   R509_000_POS : ALIAS FOR R509[0].POS;
   R6 : CONTROL[51];
   R97 : CONTROL[2] := ([0].LEN := 10, [1].LEN := 10);
        [0]   // LEHR SPEED Control word For Lehr Speed averaging Function
        [1]   // LEHR SPEED Control word For lehr Speed standard Deviation
   REL_CRUSH_ALL_OFF : ALIAS FOR I[73].10;
   REL_CRUSH_ALL_ON : ALIAS FOR I[73].11;
   REL_DATARCVD_N : ALIAS FOR O[54].2;
   REL_DATARCVDS : ALIAS FOR O[58].2;
   REL_REJWINLAMPN : ALIAS FOR O[54].3;
   REL_REJWINLAMPS : ALIAS FOR O[58].3;
   Sbr_IN_dCapIndex : DINT; {access Read Only}
   Sbr_IN_dConveyor : DINT; {access Read Only}
   Sbr_IN_dDataLength : DINT; {access Read Only}
   Sbr_IN_DestinationCullet : DINT; {access Read Only}
   Sbr_IN_DestinationID : DINT; {access Read Only}
   Sbr_IN_dIndexHead : DINT; {access Read Only}
   Sbr_IN_dMaskAllowed : DINT; {access Read Only}
   Sbr_IN_Position : DINT; {access Read Only}
   Sbr_IN_PosStart : DINT; {access Read Only}
   Sbr_IN_PosStop : DINT; {access Read Only}
   Sbr_IN_ReasonID : DINT; {access Read Only}
   Sbr_IN_ReentryPosition : DINT; {access Read Only}
   Sbr_IN_ReentryPosition_max : DINT; {access Read Only}
   Sbr_IN_ReentryPosition_min : DINT; {access Read Only}
   Sbr_IN_xHeadPos : BOOL; {access Read Only}
   Sbr_IN_xSendAllCullet : BOOL; {access Read Only}
   Sbr_INO_DestinationLite : DINT; {access Read Only}
   Sbr_INO_tConvoy_SL : UDT_Convoy_SL; {access Read Only}
   Sbr_INO_tConvoyCap_ZC : UDT_ConvoyCap_ZC; {access Read Only}
   Sbr_INO_xALLForDestination : BOOL; {access Read Only}
   Sbr_INO_xAllLiteToCullet : BOOL; {access Read Only}
   Sbr_INO_xAtLeastOneForDestination : BOOL; {access Read Only}
   Sbr_INO_xAtLeastOneToCullet : BOOL; {access Read Only}
   Sbr_OUT_dIndexTail : DINT; {access Read Only}
   Sbr_OUT_dTotalCaps : DINT; {access Read Only}
   Sbr_OUT_ReqRot_CCW : BOOL; {access Read Only}
   Sbr_OUT_ReqRot_CW : BOOL; {access Read Only}
   Sbr_OUT_rgdConvoyGaps : DINT[4]; {access Read Only}
   Sbr_OUT_rgdConvoyLengths : DINT[4]; {access Read Only}
   SLOW_BLINK : ALIAS FOR T4[0];
   Speed_Offset_CM07N : DINT := -20;   // This was added to allow for speed adjustment to CM07N
   Speed_Offset_Result_CM07N : DINT := 237;
   T103 : TIMER[1];
   T108 : TIMER[1];
   T113 : TIMER[1];
   T118 : TIMER[1];
   T123 : TIMER[1];
   T128 : TIMER[1];
   T133 : TIMER[1];
   T182 : TIMER[11] := ([0].PRE := 5, [0].ACC := 5, [0].EN := 1, [0].DN := 1, [1].PRE := 50, [2].PRE := 1, [2].ACC := 3, [2].EN := 1, [2].DN := 1, [3].PRE := 30, [4].PRE := 10, [5].PRE := 20000, [5].ACC := 25, [5].EN := 1, [5].TT := 1, [6].PRE := 100, [7].PRE := 500, [8].PRE := 500, [8].ACC := 201, [8].EN := 1, [8].TT := 1, [9].PRE := 10, [10].PRE := 100);
        [7]   // VMCC M2 Speed zone 2 Start Test Timer * M2CM2
        [8]   // VMCC M2 Speed zone 2 Stop Test Timer * M2CM2
   T4 : TIMER[51] := ([0].PRE := 1000, [0].ACC := 220, [0].EN := 1, [0].TT := 1, [1].PRE := 1000, [2].PRE := 500, [3].PRE := 500, [4].PRE := 10000, [8].PRE := 200, [9].PRE := 500, [10].PRE := 500, [11].PRE := 60, [13].PRE := 60000, [13].ACC := 60002, [13].EN := 1, [13].DN := 1, [26].PRE := 2500, [27].PRE := 2500, [28].PRE := 2500, [29].PRE := 2500, [30].PRE := 12000, [30].ACC := 12001, [30].EN := 1, [30].DN := 1, [31].PRE := 100, [31].ACC := 101, [31].EN := 1, [31].DN := 1, [33].PRE := 2500, [34].PRE := 2500, [35].PRE := 2500, [36].PRE := 2500, [37].PRE := 2500, [38].PRE := 2500, [39].PRE := 2500, [40].PRE := 2500, [41].PRE := 2500, [42].PRE := 2500, [43].PRE := 2500, [44].PRE := 2500, [45].PRE := 2500, [46].PRE := 2500, [47].PRE := 2500, [48].PRE := 2500, [49].PRE := 2500, [50].PRE := 2500);
        [0]   // Slow blink On time Timer
        [44]   // M2CM09N Running Delay Timer
        [31]   // M2CMO2 Stopped Failure Detect Debounce timer
        [43]   // M2CM09S Running Delay Timer
        [42]   // M2CM08N Running Delay Timer
        [1]   // Slow blink off time timer
        [26]   // M2CM01 Running Delay Timer
        [29]   // M2CM04S Running Delay Timer
        [2]   // Fast blink On time timer
        [28]   // M2CM03 Running Delay Timer
        [3]   // Fast Blink off time timer
        [39]   // M2CM07S Running Delay Timer
        [8]   // Conv 12 drive enable timer
        [27]   // M2CM02 Running Delay Timer
        [34]   // M2CM04N Running Delay Timer
        [35]   // M2CM05S Running Delay Timer
        [38]   // M2CM06N Running Delay Timer
        [33]   // VMCC M2 Drive Fault timer hold to see if fault will clear
        [37]   // M2CM06S Running Delay Timer
        [36]   // M2CM05N Running Delay Timer
        [40]   // M2CM07N Running Delay Timer
        [41]   // M2CM08S Running Delay Timer
        [46]   // M2CM10N Running Delay Timer
        [47]   // M2CM11S Running Delay Timer
        [48]   // M2CM011N Running Delay Timer
        [49]   // M2CM012S Running Delay Timer
        [30]   // Drive Stopped Failure Detect Debounce timer (All drives were running prev)
        [13]   // BENCHBOARD Timer for CROSSBREAK ON duration (60 sec.)
        [11]   // Test Timer
        [4]   // M4-->>M2 Mainline Sec. Trans. Backup delay timer
        [50]   // M2CM012N Running Delay Timer
        [45]   // M2CM10S Running Delay Timer
   T47 : TIMER[32];
        [10]   // Conveyor 10 Resync Input Debounce Timer
        [11]   // Conveyor 11 Resync Input Debounce Timer
        [12]   // Conveyor 12 Resync Input Debounce Timer
        [19]   // Conveyor 19 Resync Input Debounce Timer
        [1]   // Conveyor 1 Resync Input Debounce Timer
        [20]   // Conveyor 20 Resync Input Debounce Timer
        [21]   // Conveyor 21 Resync Input Debounce Timer
        [22]   // Conveyor 22 Resync Input Debounce Timer
        [23]   // Conveyor 23 Resync Input Debounce Timer
        [24]   // Conveyor 24 Resync Input Debounce Timer
        [25]   // Conveyor 25 Resync Input Debounce Timer
        [26]   // Conveyor 26 Resync Input Debounce Timer
        [27]   // Conveyor 27 Resync Input Debounce Timer
        [28]   // Conveyor 28 Resync Input Debounce Timer
        [29]   // Conveyor 29 Resync Input Debounce Timer
        [2]   // Conveyor 2 Resync Input Debounce Timer
        [30]   // Conveyor 30 Resync Input Debounce Timer
        [31]   // Conveyor 31 Resync Input Debounce Timer
        [13]   // Conveyor 13 Resync Input Debounce Timer
        [3]   // Conveyor 3 Resync Input Debounce Timer
        [4]   // Conveyor 4 Resync Input Debounce Timer
        [5]   // Conveyor 5 Resync Input Debounce Timer
        [6]   // Conveyor 6 Resync Input Debounce Timer
        [7]   // Conveyor 7 Resync Input Debounce Timer
        [8]   // Conveyor 8 Resync Input Debounce Timer
        [9]   // Conveyor 9 Resync Input Debounce Timer
        [14]   // Conveyor 14 Resync Input Debounce Timer
        [15]   // Conveyor 15 Resync Input Debounce Timer
        [16]   // Conveyor 16 Resync Input Debounce Timer
        [17]   // Conveyor 17 Resync Input Debounce Timer
        [18]   // Conveyor 18 Resync Input Debounce Timer
   T9 : TIMER[22] := ([10].PRE := 8000, [10].ACC := 8002, [10].EN := 1, [10].DN := 1, [11].PRE := 8000, [11].ACC := 8001, [11].EN := 1, [11].DN := 1, [12].PRE := 8000, [12].ACC := 8001, [12].EN := 1, [12].DN := 1, [13].PRE := 8000, [13].ACC := 8002, [13].EN := 1, [13].DN := 1, [14].PRE := 8000, [14].ACC := 8001, [14].EN := 1, [14].DN := 1, [15].PRE := 8000, [15].ACC := 8000, [15].EN := 1, [15].DN := 1, [16].PRE := 8000, [16].ACC := 8002, [16].EN := 1, [16].DN := 1, [17].PRE := 8000, [17].ACC := 8002, [17].EN := 1, [17].DN := 1, [18].PRE := 8000, [18].ACC := 8001, [18].EN := 1, [18].DN := 1, [19].PRE := 8000, [19].ACC := 8000, [19].EN := 1, [19].DN := 1, [20].PRE := 8000, [20].ACC := 8001, [20].EN := 1, [20].DN := 1, [21].PRE := 8000, [21].ACC := 8001, [21].EN := 1, [21].DN := 1);
        [10]   // Conv 1 drive enable timer
        [11]   // Conv 2 drive enable timer
        [12]   // Conv 3 drive enable timer
        [13]   // Conv 4 drive enable timer
        [14]   // Conv 5 drive enable timer
        [15]   // Conv 6 drive enable timer
        [16]   // Conv 7 drive enable timer
        [17]   // Conv 8 drive enable timer
        [18]   // Conv 9 drive enable timer
        [19]   // Conv 10 drive enable timer
        [20]   // Conv 11 drive enable timer
        [21]   // Conv 12 drive enable timer
   T95 : TIMER[10] := ([0].PRE := 1000);
        [0].DN   // LEHR SPEED Sample Period timer Elapsed
        [0]   // LEHR SPEED Sample period Timer
   TD1_N_MOVIN : ALIAS FOR N14[256].2;
   TD1_N_MOVOUT : ALIAS FOR N14[257].2;
   TD1_S_MOVIN : ALIAS FOR N14[256].3;
   TD1_S_MOVOUT : ALIAS FOR N14[257].3;
   TD2_N_MOVIN : ALIAS FOR N14[256].4;
   TD2_N_MOVOUT : ALIAS FOR N14[257].4;
   TD2_S_MOVIN : ALIAS FOR N14[256].5;
   TD2_S_MOVOUT : ALIAS FOR N14[257].5;
   TD3_N_MOVIN : ALIAS FOR N14[256].6;
   TD3_N_MOVOUT : ALIAS FOR N14[257].6;
   TD3_S_MOVIN : ALIAS FOR N14[256].7;
   TD3_S_MOVOUT : ALIAS FOR N14[257].7;
   TD4_N_MOVIN : ALIAS FOR N14[256].8;
   TD4_N_MOVOUT : ALIAS FOR N14[257].8;
   TD4_S_MOVIN : ALIAS FOR N14[256].9;
   TD4_S_MOVOUT : ALIAS FOR N14[257].9;
   TD5_N_MOVIN : ALIAS FOR N14[256].10;
   TD5_N_MOVOUT : ALIAS FOR N14[257].10;
   TD5_S_MOVIN : ALIAS FOR N14[256].11;
   TD5_S_MOVOUT : ALIAS FOR N14[257].11;
   TD_ALM_HORN_RLY : ALIAS FOR O[21].3;
   TD_ALM_LAMP : ALIAS FOR I[18].4;
   TD_ALM_RESET : ALIAS FOR I[17].9;
   TD_ALM_SILENCE : ALIAS FOR I[17].8;
   TD_AMBER_STKLTE : ALIAS FOR O[21].6;
   TD_BLUE_STKLTE : ALIAS FOR O[21].5;
   TD_CS2S_Crush_All_Stacklight : ALIAS FOR O[70].15;   // Red Light mounted on the top of panel
   TD_DC_INPWR : ALIAS FOR I[17].2;
   TD_DC_OUTPWR : ALIAS FOR I[17].3;
   TD_DC_PS1 : ALIAS FOR I[17].4;
   TD_DC_PS2 : ALIAS FOR I[17].6;
   TD_DC_PS3 : ALIAS FOR I[17].7;
   TD_DRV_CONT_ON : ALIAS FOR I[17].1;
   TD_DRV_FLT_LMP : ALIAS FOR O[21].0;
   TD_ESTOP : ALIAS FOR I[17].10;
   TD_ESTOPPWR : ALIAS FOR I[17].5;
   TD_FLT_RES_RLY : ALIAS FOR O[21].1;
   TD_RED_STKLTE : ALIAS FOR O[21].4;
   TDN_CRUSH_ALL_OFF : ALIAS FOR I[44].12;
   TDN_CRUSH_ALL_ON : ALIAS FOR I[44].13;
   TDN_FLT : ALIAS FOR I[18].1;
   TDN_FWD : ALIAS FOR O[20].1;
   TDN_REV : ALIAS FOR O[20].5;
   TDN_SS1 : ALIAS FOR O[20].13;
   TDN_SS2 : ALIAS FOR O[20].9;
   TDS_CRUSH_ALL_OFF : ALIAS FOR I[64].12;
   TDS_CRUSH_ALL_ON : ALIAS FOR I[64].13;
   TDS_FLT : ALIAS FOR I[18].2;
   TDS_FWD : ALIAS FOR O[20].2;
   TDS_REV : ALIAS FOR O[20].6;
   TDS_SS1 : ALIAS FOR O[20].14;
   TDS_SS2 : ALIAS FOR O[20].10;
   TEST_OPERAND : ALIAS FOR N7[11];
   TEST_TIMER : ALIAS FOR T4[11];
   TK1_N_MOVDN : ALIAS FOR N14[253].2;
   TK1_N_MOVIN : ALIAS FOR N14[254].2;
   TK1_N_MOVOUT : ALIAS FOR N14[255].2;
   TK1_N_MOVUP : ALIAS FOR N14[252].2;
   TK1_S_MOVDN : ALIAS FOR N14[253].3;
   TK1_S_MOVIN : ALIAS FOR N14[254].3;
   TK1_S_MOVOUT : ALIAS FOR N14[255].3;
   TK1_S_MOVUP : ALIAS FOR N14[252].3;
   TK2_N_MOVDN : ALIAS FOR N14[253].4;
   TK2_N_MOVIN : ALIAS FOR N14[254].4;
   TK2_N_MOVOUT : ALIAS FOR N14[255].4;
   TK2_N_MOVUP : ALIAS FOR N14[252].4;
   TK2_S_MOVDN : ALIAS FOR N14[253].5;
   TK2_S_MOVIN : ALIAS FOR N14[254].5;
   TK2_S_MOVOUT : ALIAS FOR N14[255].5;
   TK2_S_MOVUP : ALIAS FOR N14[252].5;
   TK3_N_MOVDN : ALIAS FOR N14[253].6;
   TK3_N_MOVIN : ALIAS FOR N14[254].6;
   TK3_N_MOVOUT : ALIAS FOR N14[255].6;
   TK3_N_MOVUP : ALIAS FOR N14[252].6;
   TK3_S_MOVDN : ALIAS FOR N14[253].7;
   TK3_S_MOVIN : ALIAS FOR N14[254].7;
   TK3_S_MOVOUT : ALIAS FOR N14[255].7;
   TK3_S_MOVUP : ALIAS FOR N14[252].7;
   TK4_N_MOVDN : ALIAS FOR N14[253].8;
   TK4_N_MOVIN : ALIAS FOR N14[254].8;
   TK4_N_MOVOUT : ALIAS FOR N14[255].8;
   TK4_N_MOVUP : ALIAS FOR N14[252].8;
   TK4_S_MOVDN : ALIAS FOR N14[253].9;
   TK4_S_MOVIN : ALIAS FOR N14[254].9;
   TK4_S_MOVOUT : ALIAS FOR N14[255].9;
   TK4_S_MOVUP : ALIAS FOR N14[252].9;
   TK5_N_MOVDN : ALIAS FOR N14[253].10;
   TK5_N_MOVIN : ALIAS FOR N14[254].10;
   TK5_N_MOVOUT : ALIAS FOR N14[255].10;
   TK5_N_MOVUP : ALIAS FOR N14[252].10;
   TK5_S_MOVDN : ALIAS FOR N14[253].11;
   TK5_S_MOVIN : ALIAS FOR N14[254].11;
   TK5_S_MOVOUT : ALIAS FOR N14[255].11;
   TK5_S_MOVUP : ALIAS FOR N14[252].11;
   TK_FLT : ALIAS FOR I[18].0;
   TK_FWD : ALIAS FOR O[20].0;
   TK_REV : ALIAS FOR O[20].4;
   TK_SS1 : ALIAS FOR O[20].12;
   TK_SS2 : ALIAS FOR O[20].8;
   TMP_CenterLites : BOOL; {access Read Only}
   TMP_d : DINT; {access Read Only}
   TMP_d2 : DINT; {access Read Only}
   TMP_dAccSpace : DINT; {access Read Only}
   TMP_dActualOnLHS : DINT; {access Read Only}
   TMP_dActualSpeed : DINT; {access Read Only}
   TMP_dALARM_RT999 : DINT := 9999; {access None}
   TMP_dBaryc_ins_max : DINT; {access Read Only}
   TMP_dBaryc_ins_min : DINT; {access Read Only}
   TMP_dBufferIndex : DINT; {access Read Only}
   TMP_dBufferSize : DINT; {access Read Only}
   TMP_dCap : DINT; {access Read Only}
   TMP_dCapNextConvoy : DINT; {access Read Only}
   TMP_dConv : DINT; {access Read Only}
   TMP_dConvDebug : DINT; {access Read Only}
   TMP_dConveyorLength : DINT; {access Read Only}
   TMP_dConveyorNumberForZoneCleaning : DINT; {access Read Only}
   TMP_dConvoySearchMax : DINT; {access Read Only}
   TMP_dCountDest : DINT; {access Read Only}
   TMP_dCulletMask : DINT; {access Read Only}
   TMP_dDebug : DINT; {access Read Only}
   TMP_dDecelerationPositionEndConveyor : DINT; {access Read Only}
   TMP_dDecSpace : DINT; {access Read Only}
   TMP_dDestFile : DINT := 205; {access None}
   TMP_dDestOffset : DINT := 1; {access None}
   TMP_dDiffPhotocellStartConv0 : DINT; {access Read Only}
   TMP_dDirection : DINT; {access None}
   TMP_dEndConveyorPos : DINT; {access Read Only}
   TMP_dEndSearch0 : DINT; {access Read Only}
   TMP_dEndSearch1 : DINT; {access Read Only}
   TMP_dErrDestFile : DINT; {access None}
   TMP_dErrSourceFile : DINT; {access None}
   TMP_dFixedSideOffset : DINT; {access Read Only}
   TMP_dFixedSideOffsetBoth : DINT; {access Read Only}
   TMP_dFixedSideOffsetConvoy : DINT; {access Read Only}
   TMP_dFixedSideOffsetDW : DINT; {access Read Only}
   TMP_dFixedSideOffsetUP : DINT; {access Read Only}
   TMP_dHalfConveyorLength : DINT; {access Read Only}
   TMP_dHalfPlateLength : DINT; {access Read Only}
   TMP_dHalfWidthDifference : DINT; {access Read Only}
   TMP_dHeadMax : DINT; {access Read Only}
   TMP_dHeadPosition : DINT; {access Read Only}
   TMP_dHeadPosition_mm : DINT; {access Read Only}
   TMP_dIndC : DINT; {access Read Only}
   TMP_dIndex : DINT := 200;
   TMP_dIndex2 : DINT; {access Read Only}
   TMP_dIndex3 : DINT; {access Read Only}
   TMP_dIndex4 : DINT; {access Read Only}
   TMP_dIndexCap : DINT; {access Read Only}
   TMP_dIndexCapConv : DINT; {access Read Only}
   TMP_dIndexConv : DINT; {access Read Only}
   TMP_dIndexMotor : DINT; {access Read Only}
   TMP_dIndexNext : DINT; {access Read Only}
   TMP_dIndexNextDebug : DINT; {access Read Only}
   TMP_dIndexPlate : DINT; {access Read Only}
   TMP_dIndexPrevious : DINT; {access Read Only}
   TMP_dIndexPreviousDebug : DINT; {access Read Only}
   TMP_DistanceLateralSquaringToCenter : DINT; {access Read Only}
   TMP_dLastConv : DINT; {access Read Only}
   TMP_dLastConvTail : DINT; {access Read Only}
   TMP_dLehrSpeed : DINT; {access Read Only}
   TMP_dLineSize : DINT; {access Read Only}
   TMP_dLineSpeed : DINT; {access Read Only}
   TMP_dLite : DINT; {access Read Only}
   TMP_dLiteInv : DINT; {access Read Only}
   TMP_dManualTargetPos : DINT; {access Read Only}
   TMP_dMask : DINT; {access Read Only}
   TMP_dMaskAllowed : DINT; {access Read Only}
   TMP_dMaxCap : DINT; {access Read Only}
   TMP_dMaxLite : DINT; {access Read Only}
   TMP_dMinTail : DINT; {access Read Only}
   TMP_dMissingOnLHS : DINT; {access Read Only}
   TMP_dNextCap : DINT; {access Read Only}
   TMP_dNumFile : DINT := 648; {access None}
   TMP_dNumValues : DINT := 99; {access None}
   TMP_dOffset : DINT := 32; {access None}
   TMP_dOffsetLoadUnload_cmm : DINT; {access Read Only}
   TMP_dPhEndPosition_cmm : DINT; {access Read Only}
   TMP_dPointer : DINT; {access Read Only}
   TMP_dPointerCap : DINT; {access Read Only}
   TMP_dPos_cmm : DINT; {access Read Only}
   TMP_dPosHead_cmm : DINT; {access Read Only}
   TMP_dPosTail_cmm : DINT; {access Read Only}
   TMP_dRampMotor : DINT; {access Read Only}
   TMP_dSourceFile : DINT := 200; {access None}
   TMP_dSourceOffset : DINT; {access None}
   TMP_dStart0 : DINT; {access Read Only}
   TMP_dStart1 : DINT; {access Read Only}
   TMP_dStartSearch : DINT; {access Read Only}
   TMP_dStartSearch0 : DINT; {access Read Only}
   TMP_dStartSearch1 : DINT; {access Read Only}
   TMP_dStartSearchStop : DINT; {access Read Only}
   TMP_dStepAdvMotor : DINT; {access Read Only}
   TMP_dStop0 : DINT; {access Read Only}
   TMP_dStop1 : DINT; {access Read Only}
   TMP_dStopSearch : DINT; {access Read Only}
   TMP_dStopSearchStop : DINT; {access Read Only}
   TMP_dTailOnNextConveyor_cmm : DINT; {access Read Only}
   TMP_dTailPosition : DINT; {access Read Only}
   TMP_dTarget : DINT := 1815; {access None}
   TMP_dTotalLength : DINT; {access Read Only}
   TMP_dWander : DINT; {access Read Only}
   TMP_dWidth_mm : DINT; {access Read Only}
   TMP_HeadPos : DINT; {access Read Only}
   TMP_IdxLite : DINT; {access Read Only}
   TMP_LiteAHeadY : DINT; {access Read Only}
   TMP_LiteATailY : DINT; {access Read Only}
   TMP_LiteBHeadY : DINT; {access Read Only}
   TMP_LiteBTailY : DINT; {access Read Only}
   TMP_MOV_dDestinationVar_1 : DINT := 205; {access None}
   TMP_MOV_dDestinationVar_2 : DINT; {access None}
   TMP_MOV_dSource : DINT; {access None}
   TMP_OUT_xPlateEndTracking : BOOL; {access Read Only}
   TMP_Portrait : BOOL; {access Read Only}
   TMP_r : REAL; {access Read Only}
   TMP_r1 : REAL := 1900.0; {access None}
   TMP_rAcc : REAL := 1200.0; {access None}
   TMP_rActualValue_cmm : REAL; {access Read Only}
   TMP_rDec : REAL := 1200.0; {access None}
   TMP_rgdIndexC : DINT[4] := ([0] := 2); {access None}
   TMP_rgdPnt : DINT[5]; {access Read Only}
   TMP_rgxId : DINT[10]; {access Read Only}
   TMP_rSpeed : REAL := 1500.0; {access None}
   TMP_rTarget : REAL; {access Read Only}
   TMP_rTarget_M1 : REAL; {access Read Only}
   TMP_rTarget_M2 : REAL; {access Read Only}
   TMP_rTarget_M3 : REAL; {access Read Only}
   TMP_SendToCullet : BOOL; {access Read Only}
   TMP_SquaringPosition : DINT; {access Read Only}
   TMP_StartPlusLength : DINT; {access Read Only}
   TMP_string : STRING; {access Read Only}
   TMP_x : BOOL; {access Read Only}
   TMP_xAllCullet : BOOL; {access Read Only}
   TMP_xALLForSideLeg : BOOL; {access Read Only}
   TMP_xAllLiteToCullet : BOOL; {access Read Only}
   TMP_xAlwaysOFF : BOOL; {access Read Only}
   TMP_xAtLeastOneForQuality : BOOL; {access Read Only}
   TMP_xAtLeastOneForSideLeg : BOOL; {access Read Only}
   TMP_xAtLeastOneOK : BOOL; {access Read Only}
   TMP_xAtLeastOneToCullet : BOOL; {access Read Only}
   TMP_xCenterFound : BOOL; {access Read Only}
   TMP_xConveyorInvolvedInCleaning : BOOL; {access Read Only}
   TMP_xConveyorOfStartCleaning : BOOL; {access Read Only}
   TMP_xCulletPresent : BOOL; {access Read Only}
   TMP_xDebugOFF : BOOL; {access Read Only}
   TMP_xDebugON : BOOL := 1; {access Read Only}
   TMP_xDummy : BOOL; {access Read Only}
   TMP_xEnableLoadUnload : BOOL; {access Read Only}
   TMP_xEnableZoneCleaning : BOOL; {access Read Only}
   TMP_xFirstConv : BOOL; {access Read Only}
   TMP_xForwardCommadnForCleaningZone : BOOL; {access Read Only}
   TMP_xInitialize : BOOL; {access None}
   TMP_xJustOnePlateMissing : BOOL; {access Read Only}
   TMP_xLastConv : BOOL; {access Read Only}
   TMP_xLastConvDebug : BOOL; {access Read Only}
   TMP_xLastModalityLoadBwd : BOOL; {access Read Only}
   TMP_xLastModalityUnloadBwd : BOOL; {access Read Only}
   TMP_xLiteThisDestPresent : BOOL; {access Read Only}
   TMP_xMinTailFound : BOOL; {access Read Only}
   TMP_xOSN : DINT; {access None}
   TMP_xOSN_B : DINT; {access Read Only}
   TMP_xOSR : DINT; {access None}
   TMP_xOSR_B : DINT; {access Read Only}
   TMP_xOSRDebug : BOOL := 1; {access Read Only}
   TMP_xPlateFound : BOOL; {access Read Only}
   TMP_xPlateOnConvoyOnNextConveyor : BOOL; {access Read Only}
   TMP_xPosHead : BOOL; {access Read Only}
   TMP_xPositioning : BOOL; {access Read Only}
   TMP_xPositioning_M1 : BOOL; {access Read Only}
   TMP_xPositioning_M2 : BOOL; {access Read Only}
   TMP_xPositioning_M3 : BOOL; {access Read Only}
   TMP_xPowerSaving : BOOL; {access Read Only}
   TMP_xPresenceAlternative : BOOL; {access Read Only}
   TMP_xPresenceDestination : BOOL; {access Read Only}
   TMP_xPresenceSecondDestination : BOOL; {access Read Only}
   TMP_xReqStopM310M1 : BOOL; {access Read Only}
   TMP_xReqStopM310M2 : BOOL; {access Read Only}
   TMP_xReqStopM310M3 : BOOL; {access Read Only}
   TMP_xReqStopM315M1 : BOOL; {access Read Only}
   TMP_xReqStopM315M2 : BOOL; {access Read Only}
   TMP_xReqStopM315M3 : BOOL; {access Read Only}
   TMP_xReqUnpack : BOOL; {access Read Only}
   TMP_xReverse : BOOL; {access Read Only}
   TMP_xReverse_M1 : BOOL; {access Read Only}
   TMP_xReverse_M2 : BOOL; {access Read Only}
   TMP_xReverse_M3 : BOOL; {access Read Only}
   TMP_xRun : BOOL; {access Read Only}
   TMP_xRun_M1 : BOOL; {access Read Only}
   TMP_xRun_M2 : BOOL; {access Read Only}
   TMP_xRun_M3 : BOOL; {access Read Only}
   TMP_xSimulationActive : BOOL; {access Read Only}
   TMP_xTailFound : BOOL; {access Read Only}
   TMP_xYInversionLite : BOOL; {access Read Only}
   TMP_xYWithBarycenter : BOOL; {access Read Only}
   TMR_Power_Cycle : TIMER := (PRE := 1000, ACC := 1001, EN := 1, DN := 1);
   tony_always_false : BOOL; {access Read Only}
   TRIM_SPEED : ALIAS FOR N20[2];
   TZ1_K_NTH_ADJ : ALIAS FOR O[19].2;
   TZ1_K_STH_ADJ : ALIAS FOR O[19].3;
   TZ1_N_AUTO : ALIAS FOR N14[250].2;
   TZ1_N_MANL : ALIAS FOR N14[251].2;
   TZ1_S_AUTO : ALIAS FOR N14[250].3;
   TZ1_S_MANL : ALIAS FOR N14[251].3;
   TZ1_T_NTH_ADJ : ALIAS FOR O[22].2;
   TZ1_T_STH_ADJ : ALIAS FOR O[22].3;
   TZ2_K_NTH_ADJ : ALIAS FOR O[19].4;
   TZ2_K_STH_ADJ : ALIAS FOR O[19].5;
   TZ2_N_AUTO : ALIAS FOR N14[250].4;
   TZ2_N_MANL : ALIAS FOR N14[251].4;
   TZ2_S_AUTO : ALIAS FOR N14[250].5;
   TZ2_S_MANL : ALIAS FOR N14[251].5;
   TZ2_T_NTH_ADJ : ALIAS FOR O[22].4;
   TZ2_T_STH_ADJ : ALIAS FOR O[22].5;
   TZ3_K_NTH_ADJ : ALIAS FOR O[19].6;
   TZ3_K_STH_ADJ : ALIAS FOR O[19].7;
   TZ3_N_AUTO : ALIAS FOR N14[250].6;
   TZ3_N_MANL : ALIAS FOR N14[251].6;
   TZ3_S_AUTO : ALIAS FOR N14[250].7;
   TZ3_S_MANL : ALIAS FOR N14[251].7;
   TZ3_T_NTH_ADJ : ALIAS FOR O[22].6;
   TZ3_T_STH_ADJ : ALIAS FOR O[22].7;
   TZ4_K_NTH_ADJ : ALIAS FOR O[19].8;
   TZ4_K_STH_ADJ : ALIAS FOR O[19].9;
   TZ4_N_AUTO : ALIAS FOR N14[250].8;
   TZ4_N_MANL : ALIAS FOR N14[251].8;
   TZ4_S_AUTO : ALIAS FOR N14[250].9;
   TZ4_S_MANL : ALIAS FOR N14[251].9;
   TZ4_T_NTH_ADJ : ALIAS FOR O[22].8;
   TZ4_T_STH_ADJ : ALIAS FOR O[22].9;
   TZ5_K_NTH_ADJ : ALIAS FOR O[19].10;
   TZ5_K_STH_ADJ : ALIAS FOR O[19].11;
   TZ5_N_AUTO : ALIAS FOR N14[250].10;
   TZ5_N_MANL : ALIAS FOR N14[251].10;
   TZ5_S_AUTO : ALIAS FOR N14[250].11;
   TZ5_S_MANL : ALIAS FOR N14[251].11;
   TZ5_T_NTH_ADJ : ALIAS FOR O[22].10;
   TZ5_T_STH_ADJ : ALIAS FOR O[22].11;
   VIN_A_INSP_S1 : ALIAS FOR N26[30].0;
   VIN_A_INSP_S11 : ALIAS FOR N26[30].0;
   VIN_A_INSP_S2 : ALIAS FOR N26[30].1;
   VIN_A_INSP_S3 : ALIAS FOR N26[30].2;
   VIN_A_INSP_S4 : ALIAS FOR N26[30].3;
   VIN_A_INSP_S5 : ALIAS FOR N26[30].4;
   VIN_A_INSP_S6 : ALIAS FOR N26[30].5;
   VIN_A_INSP_S7 : ALIAS FOR N26[30].6;
   VIN_A_INSP_S8 : ALIAS FOR N26[30].7;
   VIN_A_INSP_S9 : ALIAS FOR N26[30].8;
   VIN_A_INSP_WD : ALIAS FOR N26[30];
   VIN_B_INSP_S1 : ALIAS FOR N26[31].0;
   VIN_B_INSP_S2 : ALIAS FOR N26[31].1;
   VIN_B_INSP_S3 : ALIAS FOR N26[31].2;
   VIN_B_INSP_S4 : ALIAS FOR N26[31].3;
   VIN_B_INSP_S5 : ALIAS FOR N26[31].4;
   VIN_B_INSP_S6 : ALIAS FOR N26[31].5;
   VIN_B_INSP_S7 : ALIAS FOR N26[31].6;
   VIN_B_INSP_S8 : ALIAS FOR N26[31].7;
   VIN_B_INSP_S9 : ALIAS FOR N26[31].8;
   VIN_B_INSP_WD : ALIAS FOR N26[31];
   VIN_C_INSP_S1 : ALIAS FOR N26[32].0;
   VIN_C_INSP_S2 : ALIAS FOR N26[32].1;
   VIN_C_INSP_S3 : ALIAS FOR N26[32].2;
   VIN_C_INSP_S4 : ALIAS FOR N26[32].3;
   VIN_C_INSP_S5 : ALIAS FOR N26[32].4;
   VIN_C_INSP_S6 : ALIAS FOR N26[32].5;
   VIN_C_INSP_S7 : ALIAS FOR N26[32].6;
   VIN_C_INSP_S8 : ALIAS FOR N26[32].7;
   VIN_C_INSP_S9 : ALIAS FOR N26[32].8;
   VIN_C_INSP_WD : ALIAS FOR N26[32];
   VIN_D_INSP_S1 : ALIAS FOR N26[33].0;
   VIN_D_INSP_S2 : ALIAS FOR N26[33].1;
   VIN_D_INSP_S3 : ALIAS FOR N26[33].2;
   VIN_D_INSP_S4 : ALIAS FOR N26[33].3;
   VIN_D_INSP_S5 : ALIAS FOR N26[33].4;
   VIN_D_INSP_S6 : ALIAS FOR N26[33].5;
   VIN_D_INSP_S7 : ALIAS FOR N26[33].6;
   VIN_D_INSP_S8 : ALIAS FOR N26[33].7;
   VIN_D_INSP_S9 : ALIAS FOR N26[33].8;
   VIN_D_INSP_WD : ALIAS FOR N26[33];
   VIN_GRP_ID : ALIAS FOR N26[0];
   VIN_GRP_ID1 : ALIAS FOR N26[0];
   VIN_LEN_S1 : ALIAS FOR N26[21];
   VIN_LEN_S11 : ALIAS FOR N26[21];
   VIN_LEN_S2 : ALIAS FOR N26[22];
   VIN_LEN_S3 : ALIAS FOR N26[23];
   VIN_LEN_S4 : ALIAS FOR N26[24];
   VIN_LEN_S5 : ALIAS FOR N26[25];
   VIN_LEN_S6 : ALIAS FOR N26[26];
   VIN_LEN_S7 : ALIAS FOR N26[27];
   VIN_LEN_S8 : ALIAS FOR N26[28];
   VIN_LEN_S9 : ALIAS FOR N26[29];
   VIN_NTOL_CRN : ALIAS FOR N26[16];
   VIN_NTOL_EDG : ALIAS FOR N26[15];
   VIN_NTOL_LEN : ALIAS FOR N26[12];
   VIN_NTOL_SKW : ALIAS FOR N26[13];
   VIN_NTOL_SQR : ALIAS FOR N26[14];
   VIN_NTOL_WID : ALIAS FOR N26[11];
   VIN_NTOL_WID1 : ALIAS FOR N26[11];
   VIN_NUM_SPLITS : ALIAS FOR N26[4];
   VIN_NUM_SPLITS1 : ALIAS FOR N26[4];
   VIN_NUM_STRMS : ALIAS FOR N26[3];
   VIN_NUM_STRMS1 : ALIAS FOR N26[3];
   VIN_PTOL_CRN : ALIAS FOR N26[10];
   VIN_PTOL_EDG : ALIAS FOR N26[9];
   VIN_PTOL_LEN : ALIAS FOR N26[6];
   VIN_PTOL_SKW : ALIAS FOR N26[7];
   VIN_PTOL_SQR : ALIAS FOR N26[8];
   VIN_PTOL_WID : ALIAS FOR N26[5];
   VIN_PTOL_WID1 : ALIAS FOR N26[5];
   VIN_QUALITY_S1 : ALIAS FOR N26[34];
   VIN_QUALITY_S2 : ALIAS FOR N26[35];
   VIN_QUALITY_S3 : ALIAS FOR N26[36];
   VIN_QUALITY_S4 : ALIAS FOR N26[37];
   VIN_QUALITY_S5 : ALIAS FOR N26[38];
   VIN_QUALITY_S6 : ALIAS FOR N26[39];
   VIN_QUALITY_S7 : ALIAS FOR N26[40];
   VIN_QUALITY_S8 : ALIAS FOR N26[41];
   VIN_QUALITY_S9 : ALIAS FOR N26[42];
   VIN_SUB_THICK : ALIAS FOR N26[2];
   VIN_SUB_THICK1 : ALIAS FOR N26[2];
   VIN_SUB_TYPE : ALIAS FOR N26[1];
   VIN_SUB_TYPE1 : ALIAS FOR N26[1];
   VIN_WID_A : ALIAS FOR N26[17];
   VIN_WID_A1 : ALIAS FOR N26[17];
   VIN_WID_B : ALIAS FOR N26[18];
   VIN_WID_C : ALIAS FOR N26[19];
   VIN_WID_D : ALIAS FOR N26[20];
   VIS_BLUE_STACK : ALIAS FOR O[36].15;
   VIS_HB : ALIAS FOR N27[60].0;
   VIS_IGNORE_LEN_EN : ALIAS FOR N26[100].12;
   VIS_OUTPT_OFF : ALIAS FOR N27[60].2;
   VIS_PLC_RD_ERR : ALIAS FOR N27[60].3;
   VIS_SYS_STOPPED : ALIAS FOR N27[60].1;
   VISCOM_BAD : ALIAS FOR N21[3].1;
   VISCOM_ENABLE : ALIAS FOR N17[11].1;
   VISCOM_GOOD : ALIAS FOR N21[3].0;
   VISCOM_NEWLEN : ALIAS FOR N21[1];
   VISCOM_NEWWID : ALIAS FOR N21[2];
   VISCOM_RESULT : ALIAS FOR N21[3];
   VISCOM_WAIT : ALIAS FOR N17[11].0;
   VISCOMM_NEWDATA : ALIAS FOR N21[0].1;
   VOUT_GRP_ID : ALIAS FOR N27[0];
   VOUT_NEW_DATA : ALIAS FOR N27[2];
   VOUT_NUM_SPLITS : ALIAS FOR N27[4];
   VOUT_NUM_STRMS : ALIAS FOR N27[3];
   VOUT_ONLINE : ALIAS FOR N27[1].0;
   VOUT_REJ_1A : ALIAS FOR N27[5];
   VOUT_REJ_1B : ALIAS FOR N27[6];
   VOUT_REJ_1C : ALIAS FOR N27[7];
   VOUT_REJ_1D : ALIAS FOR N27[8];
   VOUT_REJ_2A : ALIAS FOR N27[9];
   VOUT_REJ_2B : ALIAS FOR N27[10];
   VOUT_REJ_2C : ALIAS FOR N27[11];
   VOUT_REJ_2D : ALIAS FOR N27[12];
   VOUT_REJ_3A : ALIAS FOR N27[13];
   VOUT_REJ_3B : ALIAS FOR N27[14];
   VOUT_REJ_3C : ALIAS FOR N27[15];
   VOUT_REJ_3D : ALIAS FOR N27[16];
   VOUT_REJ_4A : ALIAS FOR N27[17];
   VOUT_REJ_4B : ALIAS FOR N27[18];
   VOUT_REJ_4C : ALIAS FOR N27[19];
   VOUT_REJ_4D : ALIAS FOR N27[20];
   VOUT_REJ_5A : ALIAS FOR N27[21];
   VOUT_REJ_5B : ALIAS FOR N27[22];
   VOUT_REJ_5C : ALIAS FOR N27[23];
   VOUT_REJ_5D : ALIAS FOR N27[24];
   VOUT_REJ_6A : ALIAS FOR N27[25];
   VOUT_REJ_6B : ALIAS FOR N27[26];
   VOUT_REJ_6C : ALIAS FOR N27[27];
   VOUT_REJ_6D : ALIAS FOR N27[28];
   VOUT_REJ_7A : ALIAS FOR N27[29];
   VOUT_REJ_7B : ALIAS FOR N27[30];
   VOUT_REJ_7C : ALIAS FOR N27[31];
   VOUT_REJ_7D : ALIAS FOR N27[32];
   VOUT_REJ_8A : ALIAS FOR N27[33];
   VOUT_REJ_8B : ALIAS FOR N27[34];
   VOUT_REJ_8C : ALIAS FOR N27[35];
   VOUT_REJ_8D : ALIAS FOR N27[36];
   VOUT_REJ_9A : ALIAS FOR N27[37];
   VOUT_REJ_9B : ALIAS FOR N27[38];
   VOUT_REJ_9C : ALIAS FOR N27[39];
   VOUT_REJ_9D : ALIAS FOR N27[40];
   VOUT_SERV_REQ : ALIAS FOR N27[1].1;
   VOUT_STATUS : ALIAS FOR N27[1];
   VRES_GRP_ID : ALIAS FOR N25[0];
   VRES_NEW_DATA : ALIAS FOR N25[2];
   VRES_NUM_SPLITS : ALIAS FOR N25[4];
   VRES_NUM_STRMS : ALIAS FOR N25[3];
   VRES_ONLINE : ALIAS FOR N25[1].0;
   VRES_REJ_1A : ALIAS FOR N25[5];
   VRES_REJ_1B : ALIAS FOR N25[6];
   VRES_REJ_1C : ALIAS FOR N25[7];
   VRES_REJ_1D : ALIAS FOR N25[8];
   VRES_REJ_2A : ALIAS FOR N25[9];
   VRES_REJ_2B : ALIAS FOR N25[10];
   VRES_REJ_2C : ALIAS FOR N25[11];
   VRES_REJ_2D : ALIAS FOR N25[12];
   VRES_REJ_3A : ALIAS FOR N25[13];
   VRES_REJ_3B : ALIAS FOR N25[14];
   VRES_REJ_3C : ALIAS FOR N25[15];
   VRES_REJ_3D : ALIAS FOR N25[16];
   VRES_REJ_4A : ALIAS FOR N25[17];
   VRES_REJ_4B : ALIAS FOR N25[18];
   VRES_REJ_4C : ALIAS FOR N25[19];
   VRES_REJ_4D : ALIAS FOR N25[20];
   VRES_REJ_5A : ALIAS FOR N25[21];
   VRES_REJ_5B : ALIAS FOR N25[22];
   VRES_REJ_5C : ALIAS FOR N25[23];
   VRES_REJ_5D : ALIAS FOR N25[24];
   VRES_REJ_6A : ALIAS FOR N25[25];
   VRES_REJ_6B : ALIAS FOR N25[26];
   VRES_REJ_6C : ALIAS FOR N25[27];
   VRES_REJ_6D : ALIAS FOR N25[28];
   VRES_REJ_7A : ALIAS FOR N25[29];
   VRES_REJ_7B : ALIAS FOR N25[30];
   VRES_REJ_7C : ALIAS FOR N25[31];
   VRES_REJ_7D : ALIAS FOR N25[32];
   VRES_REJ_8A : ALIAS FOR N25[33];
   VRES_REJ_8B : ALIAS FOR N25[34];
   VRES_REJ_8C : ALIAS FOR N25[35];
   VRES_REJ_8D : ALIAS FOR N25[36];
   VRES_REJ_9A : ALIAS FOR N25[37];
   VRES_REJ_9B : ALIAS FOR N25[38];
   VRES_REJ_9C : ALIAS FOR N25[39];
   VRES_REJ_9D : ALIAS FOR N25[40];
   VRES_SERV_REQ : ALIAS FOR N25[1].1;
   VRES_STATUS : ALIAS FOR N25[1];
   x311PortraitMode : BOOL; {access Read Only}
   x316PortraitMode : BOOL; {access Read Only}
   xAlwaysOFF : BOOL; {access Read Only}
   xAlwaysON : BOOL := 1; {access Read Only}
   xDebugOFF : BOOL; {access Read Only}
   xDebugON : BOOL; {access Read Only}
   xSampleTablePedal : BOOL;
   Z200_SnapDataEth : UDT_ConvoyCap_ZC[2];
   Z300_BufferPlate : UDT_LINE_BUFFER_PLATE := (rgtPlate[0].tTracking.dPosition_cmm := 2872000, rgtPlate[0].tTracking.xNotConsConvTrk := 1, rgtPlate[0].tData.dLength_cmm := 90000, rgtPlate[0].tData.rgtCap[0].dConvTotLength_cmm := 90000, rgtPlate[1].tTracking.dPosition_cmm := 7466000, rgtPlate[1].tTracking.dPositionHead_cmm := 7596000, rgtPlate[1].tTracking.dPositionTail_cmm := 7336000, rgtPlate[1].tTracking.dLength_cmm := 260000, rgtPlate[1].tTracking.dIndexConvHead := 22, rgtPlate[1].tTracking.dIndexCapInConvHead := 1, rgtPlate[1].tTracking.dIndexConvTail := 21, rgtPlate[1].tTracking.dIndexCapInConvTail := 1, rgtPlate[1].tTracking.dLastConv := 22, rgtPlate[1].tTracking.dLastConvTail := 21, rgtPlate[1].tData.dLength_cmm := 260000, rgtPlate[1].tData.dTotalCaps := 1, rgtPlate[1].tData.rgtCap[0].dID := 4255229, rgtPlate[1].tData.rgtCap[0].dLength_cmm := 260000, rgtPlate[1].tData.rgtCap[0].dWidth_cmm := 360000, rgtPlate[1].tData.rgtCap[0].dThickness_cmm := 600, rgtPlate[1].tData.rgtCap[0].dGap_cmm := 30000, rgtPlate[1].tData.rgtCap[0].dFormat := 3, rgtPlate[1].tData.rgtCap[0].dNumLites := 2, rgtPlate[1].tData.rgtCap[0].dConvTotLength_cmm := 260000, rgtPlate[1].tData.rgtCap[0].dMinWidth_cmm := 360000, rgtPlate[1].tData.rgtCap[0].dMaxWidth_cmm := 360000, rgtPlate[1].tData.rgtCap[0].dGrossWidth_cmm := 377300, rgtPlate[1].tData.rgtCap[0].dDEdgeOpSide_cmm := 5000, rgtPlate[1].tData.rgtCap[0].dDEdgeOppOpSide_cmm := 5000, rgtPlate[1].tData.rgtCap[0].dCutWander_cmm := -3930, rgtPlate[1].tData.rgtCap[0].dNetWander_cmm := -6130, rgtPlate[1].tData.rgtCap[0].rgtLite[0].dID := 4255230, rgtPlate[1].tData.rgtCap[0].rgtLite[0].dProductionID := 1029, rgtPlate[1].tData.rgtCap[0].rgtLite[0].dQualityID := 10, rgtPlate[1].tData.rgtCap[0].rgtLite[0].dWidth_cmm := 180000, rgtPlate[1].tData.rgtCap[0].rgtLite[0].dBarycenter_cmm := -108930, rgtPlate[1].tData.rgtCap[0].rgtLite[1].dID := 4255231, rgtPlate[1].tData.rgtCap[0].rgtLite[1].dProductionID := 1029, rgtPlate[1].tData.rgtCap[0].rgtLite[1].dQualityID := 10, rgtPlate[1].tData.rgtCap[0].rgtLite[1].dWidth_cmm := 180000, rgtPlate[1].tData.rgtCap[0].rgtLite[1].dBarycenter_cmm := 101070, rgtPlate[1].tData.rgtCap[0].tFlag.xByYCut2 := 1, rgtPlate[1].tData.rgtCap[0].tFlag.xTrim2OpSide := 1, rgtPlate[1].tData.rgtCap[0].tFlag.xTrim1OpSide := 1, rgtPlate[1].tData.rgtCap[0].tFlag.xTrim1OppOpSide := 1, rgtPlate[1].tData.rgtCap[0].tFlag.xTrim2OppOpSide := 1, rgtPlate[1].tData.rgtCap[0].tFlag.rgxIntCut := 1, rgtPlate[1].tData.rgtCap[0].tFlag.xOptSelvedgeSel := 1, rgtPlate[1].tData.rgtCap[0].tFlag.xOptSplitBarSel := 1, rgtPlate[1].tData.rgtCap[0].tFlag.xOptSepRollSel := 1, rgtPlate[1].tData.rgtCap[0].tFlag.xHookedGeom := 1, rgtPlate[1].tData.rgtCap[0].tFlag.rgxXCutDoneHead := 2, rgtPlate[1].tData.rgtCap[0].tFlag.rgxXCutDoneTail := 2, rgtPlate[1].tData.rgtCap[0].tFlag.rgxYCutHeadDone := 835, rgtPlate[1].tData.rgtCap[0].tFlag.tSelvedgeMachine.dReqTrim2OpSide := 1, rgtPlate[1].tData.rgtCap[0].tFlag.tSelvedgeMachine.dReqTrim1OpSide := 3, rgtPlate[1].tData.rgtCap[0].tFlag.tSelvedgeMachine.dReqTrim1OppOpSide := 3, rgtPlate[1].tData.rgtCap[0].tFlag.tSelvedgeMachine.dReqTrim2OppOpSide := 1, rgtPlate[1].tData.rgtCap[0].tFlag.tSelvedgeMachine.dDoneTrim3OpSide := 3, rgtPlate[1].tData.rgtCap[0].tFlag.tSelvedgeMachine.dDoneTrim2OpSide := 1,